REGION Network 144: Change the VG2 voltage in local
   RUNG wire#powerrail
      Contact( "STATO".controllo_setVG2 )
      wire#w1
      { S7_Templates := "SrcType := Int" } GE_Contact(in1 := "STATO".stato_VOLTAGGIO_G2, in2 := 100)
      { S7_Templates := "SrcType := Int" } LE_Contact(in1 := "STATO".stato_VOLTAGGIO_G2, in2 := 1150)
      Move(in := "STATO_TMP".tmp_adj_VG2, out1 => "STATO".stato_VOLTAGGIO_G2)
      R_Coil( "STATO".controllo_setVG2 )
   END_RUNG
   RUNG wire#w1
      { S7_Templates := "SrcType := Int" } GT_Contact(in1 := "STATO".stato_VOLTAGGIO_G2, in2 := 1150)
      Move(in := 1150, out1 => "STATO".stato_VOLTAGGIO_G2)
      R_Coil( "STATO".controllo_setVG2 )
   END_RUNG
   RUNG wire#w1
      { S7_Templates := "SrcType := Int" } LT_Contact(in1 := "STATO".stato_VOLTAGGIO_G2, in2 := 100)
      Move(in := 100, out1 => "STATO".stato_VOLTAGGIO_G2)
      R_Coil( "STATO".controllo_setVG2 )
   END_RUNG
   // the same network as SCL:
   #_w1 := "STATO".controllo_setVG2 AND ("STATO".stato_VOLTAGGIO_G2 >= 100) AND ("STATO".stato_VOLTAGGIO_G2 <= 1150);
   IF #_w1 THEN "STATO".stato_VOLTAGGIO_G2 := "STATO_TMP".tmp_adj_VG2; END_IF;
   #_w2 := "STATO".controllo_setVG2;
   IF #_w1 THEN "STATO".controllo_setVG2 := FALSE; END_IF;
   #_w3 := #_w2 AND ("STATO".stato_VOLTAGGIO_G2 > 1150);
   IF #_w3 THEN
       "STATO".stato_VOLTAGGIO_G2 := 1150;
       "STATO".controllo_setVG2 := FALSE;
   END_IF;
   #_w4 := #_w2 AND ("STATO".stato_VOLTAGGIO_G2 < 100);
   IF #_w4 THEN
       "STATO".stato_VOLTAGGIO_G2 := 100;
       "STATO".controllo_setVG2 := FALSE;
   END_IF;
END_REGION

REGION Network 145: Change the VG2 voltage in remote
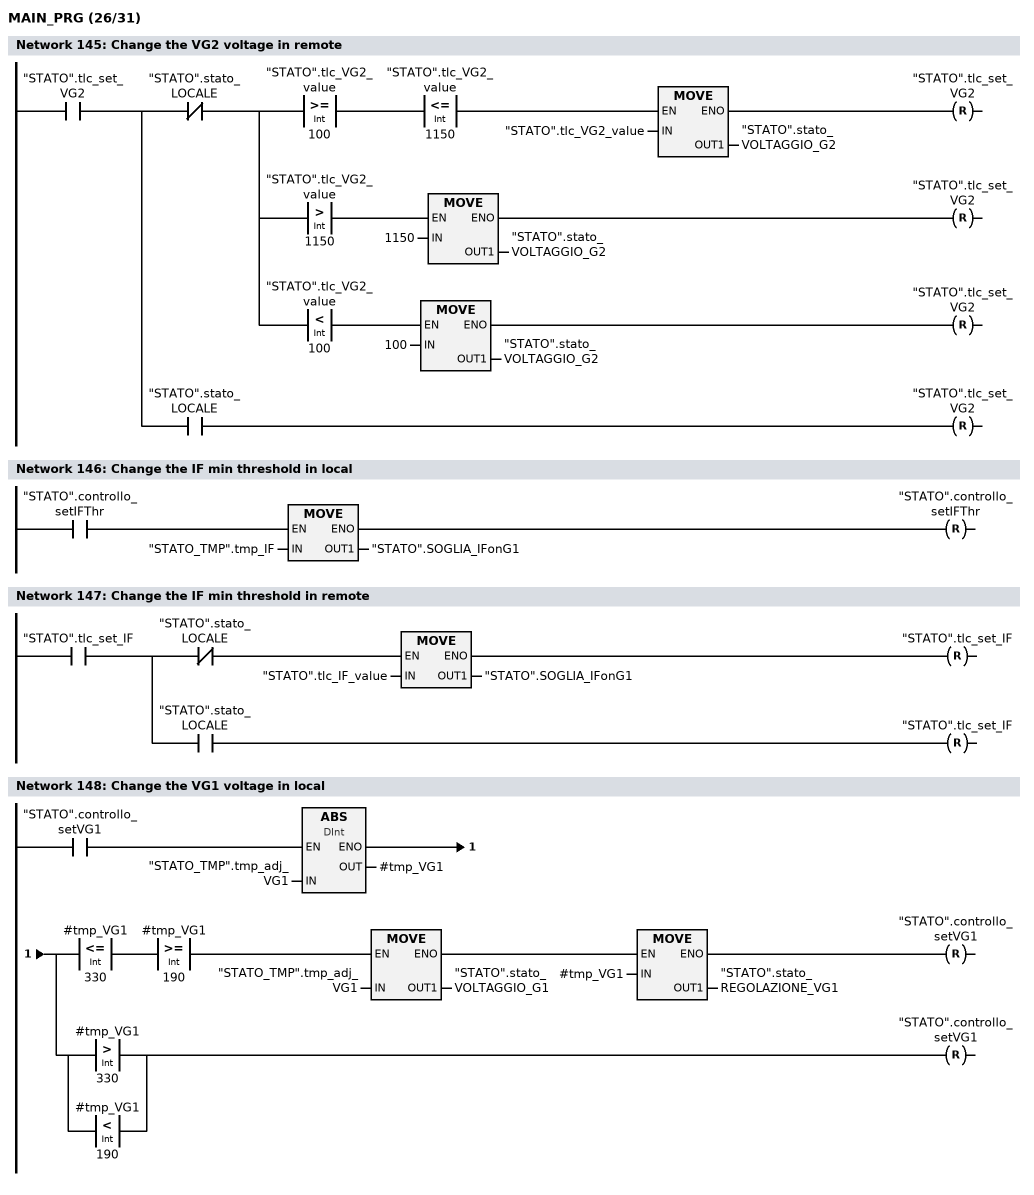
   RUNG wire#powerrail
      Contact( "STATO".tlc_set_VG2 )
      wire#w1
      I_Contact( "STATO".stato_LOCALE )
      wire#w2
      { S7_Templates := "SrcType := Int" } GE_Contact(in1 := "STATO".tlc_VG2_value, in2 := 100)
      { S7_Templates := "SrcType := Int" } LE_Contact(in1 := "STATO".tlc_VG2_value, in2 := 1150)
      Move(in := "STATO".tlc_VG2_value, out1 => "STATO".stato_VOLTAGGIO_G2)
      R_Coil( "STATO".tlc_set_VG2 )
   END_RUNG
   RUNG wire#w2
      { S7_Templates := "SrcType := Int" } GT_Contact(in1 := "STATO".tlc_VG2_value, in2 := 1150)
      Move(in := 1150, out1 => "STATO".stato_VOLTAGGIO_G2)
      R_Coil( "STATO".tlc_set_VG2 )
   END_RUNG
   RUNG wire#w2
      { S7_Templates := "SrcType := Int" } LT_Contact(in1 := "STATO".tlc_VG2_value, in2 := 100)
      Move(in := 100, out1 => "STATO".stato_VOLTAGGIO_G2)
      R_Coil( "STATO".tlc_set_VG2 )
   END_RUNG
   RUNG wire#w1
      Contact( "STATO".stato_LOCALE )
      R_Coil( "STATO".tlc_set_VG2 )
   END_RUNG
   // the same network as SCL:
   #_w1 := "STATO".tlc_set_VG2 AND NOT "STATO".stato_LOCALE;
   IF #_w1 AND ("STATO".tlc_VG2_value >= 100) AND ("STATO".tlc_VG2_value <= 1150) THEN
       "STATO".stato_VOLTAGGIO_G2 := "STATO".tlc_VG2_value;
   END_IF;
   #_w2 := "STATO".tlc_set_VG2;
   IF #_w1 AND ("STATO".tlc_VG2_value >= 100) AND ("STATO".tlc_VG2_value <= 1150) THEN
       "STATO".tlc_set_VG2 := FALSE;
   END_IF;
   IF #_w1 AND ("STATO".tlc_VG2_value > 1150) THEN
       "STATO".stato_VOLTAGGIO_G2 := 1150;
       "STATO".tlc_set_VG2 := FALSE;
   END_IF;
   IF #_w1 AND ("STATO".tlc_VG2_value < 100) THEN
       "STATO".stato_VOLTAGGIO_G2 := 100;
       "STATO".tlc_set_VG2 := FALSE;
   END_IF;
   IF #_w2 AND "STATO".stato_LOCALE THEN "STATO".tlc_set_VG2 := FALSE; END_IF;
END_REGION

REGION Network 146: Change the IF min threshold in local
   RUNG wire#powerrail
      Contact( "STATO".controllo_setIFThr )
      Move(in := "STATO_TMP".tmp_IF, out1 => "STATO".SOGLIA_IFonG1)
      R_Coil( "STATO".controllo_setIFThr )
   END_RUNG
   // the same network as SCL:
   IF "STATO".controllo_setIFThr THEN
       "STATO".SOGLIA_IFonG1 := "STATO_TMP".tmp_IF;
       "STATO".controllo_setIFThr := FALSE;
   END_IF;
END_REGION

REGION Network 147: Change the IF min threshold in remote
   RUNG wire#powerrail
      Contact( "STATO".tlc_set_IF )
      wire#w1
      I_Contact( "STATO".stato_LOCALE )
      Move(in := "STATO".tlc_IF_value, out1 => "STATO".SOGLIA_IFonG1)
      R_Coil( "STATO".tlc_set_IF )
   END_RUNG
   RUNG wire#w1
      Contact( "STATO".stato_LOCALE )
      R_Coil( "STATO".tlc_set_IF )
   END_RUNG
   // the same network as SCL:
   IF "STATO".tlc_set_IF AND NOT "STATO".stato_LOCALE THEN
       "STATO".SOGLIA_IFonG1 := "STATO".tlc_IF_value;
   END_IF;
   #_w1 := "STATO".tlc_set_IF;
   IF "STATO".tlc_set_IF AND NOT "STATO".stato_LOCALE THEN "STATO".tlc_set_IF := FALSE; END_IF;
   IF #_w1 AND "STATO".stato_LOCALE THEN "STATO".tlc_set_IF := FALSE; END_IF;
END_REGION

REGION Network 148: Change the VG1 voltage in local
   RUNG wire#powerrail
      Contact( "STATO".controllo_setVG1 )
      { S7_Templates := "SrcType := DInt" } Abs(in := "STATO_TMP".tmp_adj_VG1, out => #tmp_VG1)
      wire#w1
      { S7_Templates := "SrcType := Int" } LE_Contact(in1 := #tmp_VG1, in2 := 330)
      { S7_Templates := "SrcType := Int" } GE_Contact(in1 := #tmp_VG1, in2 := 190)
      Move(in := "STATO_TMP".tmp_adj_VG1, out1 => "STATO".stato_VOLTAGGIO_G1)
      Move(in := #tmp_VG1, out1 => "STATO".stato_REGOLAZIONE_VG1)
      R_Coil( "STATO".controllo_setVG1 )
   END_RUNG
   RUNG wire#w1
      { S7_Templates := "SrcType := Int" } GT_Contact(in1 := #tmp_VG1, in2 := 330)
      wire#w2
      R_Coil( "STATO".controllo_setVG1 )
   END_RUNG
   RUNG wire#w1
      { S7_Templates := "SrcType := Int" } LT_Contact(in1 := #tmp_VG1, in2 := 190)
   END_RUNG wire#w2
   // the same network as SCL:
   IF "STATO".controllo_setVG1 THEN #tmp_VG1 := ABS("STATO_TMP".tmp_adj_VG1); END_IF;
   IF "STATO".controllo_setVG1 AND (#tmp_VG1 <= 330) AND (#tmp_VG1 >= 190) THEN
       "STATO".stato_VOLTAGGIO_G1 := "STATO_TMP".tmp_adj_VG1;
       "STATO".stato_REGOLAZIONE_VG1 := #tmp_VG1;
   END_IF;
   #_w1 := "STATO".controllo_setVG1;
   IF "STATO".controllo_setVG1 AND (#tmp_VG1 <= 330) AND (#tmp_VG1 >= 190) THEN
       "STATO".controllo_setVG1 := FALSE;
   END_IF;
   IF #_w1 AND ((#tmp_VG1 > 330) OR (#tmp_VG1 < 190)) THEN "STATO".controllo_setVG1 := FALSE; END_IF;
END_REGION

REGION Network 149: Change the VG1 voltage in remote
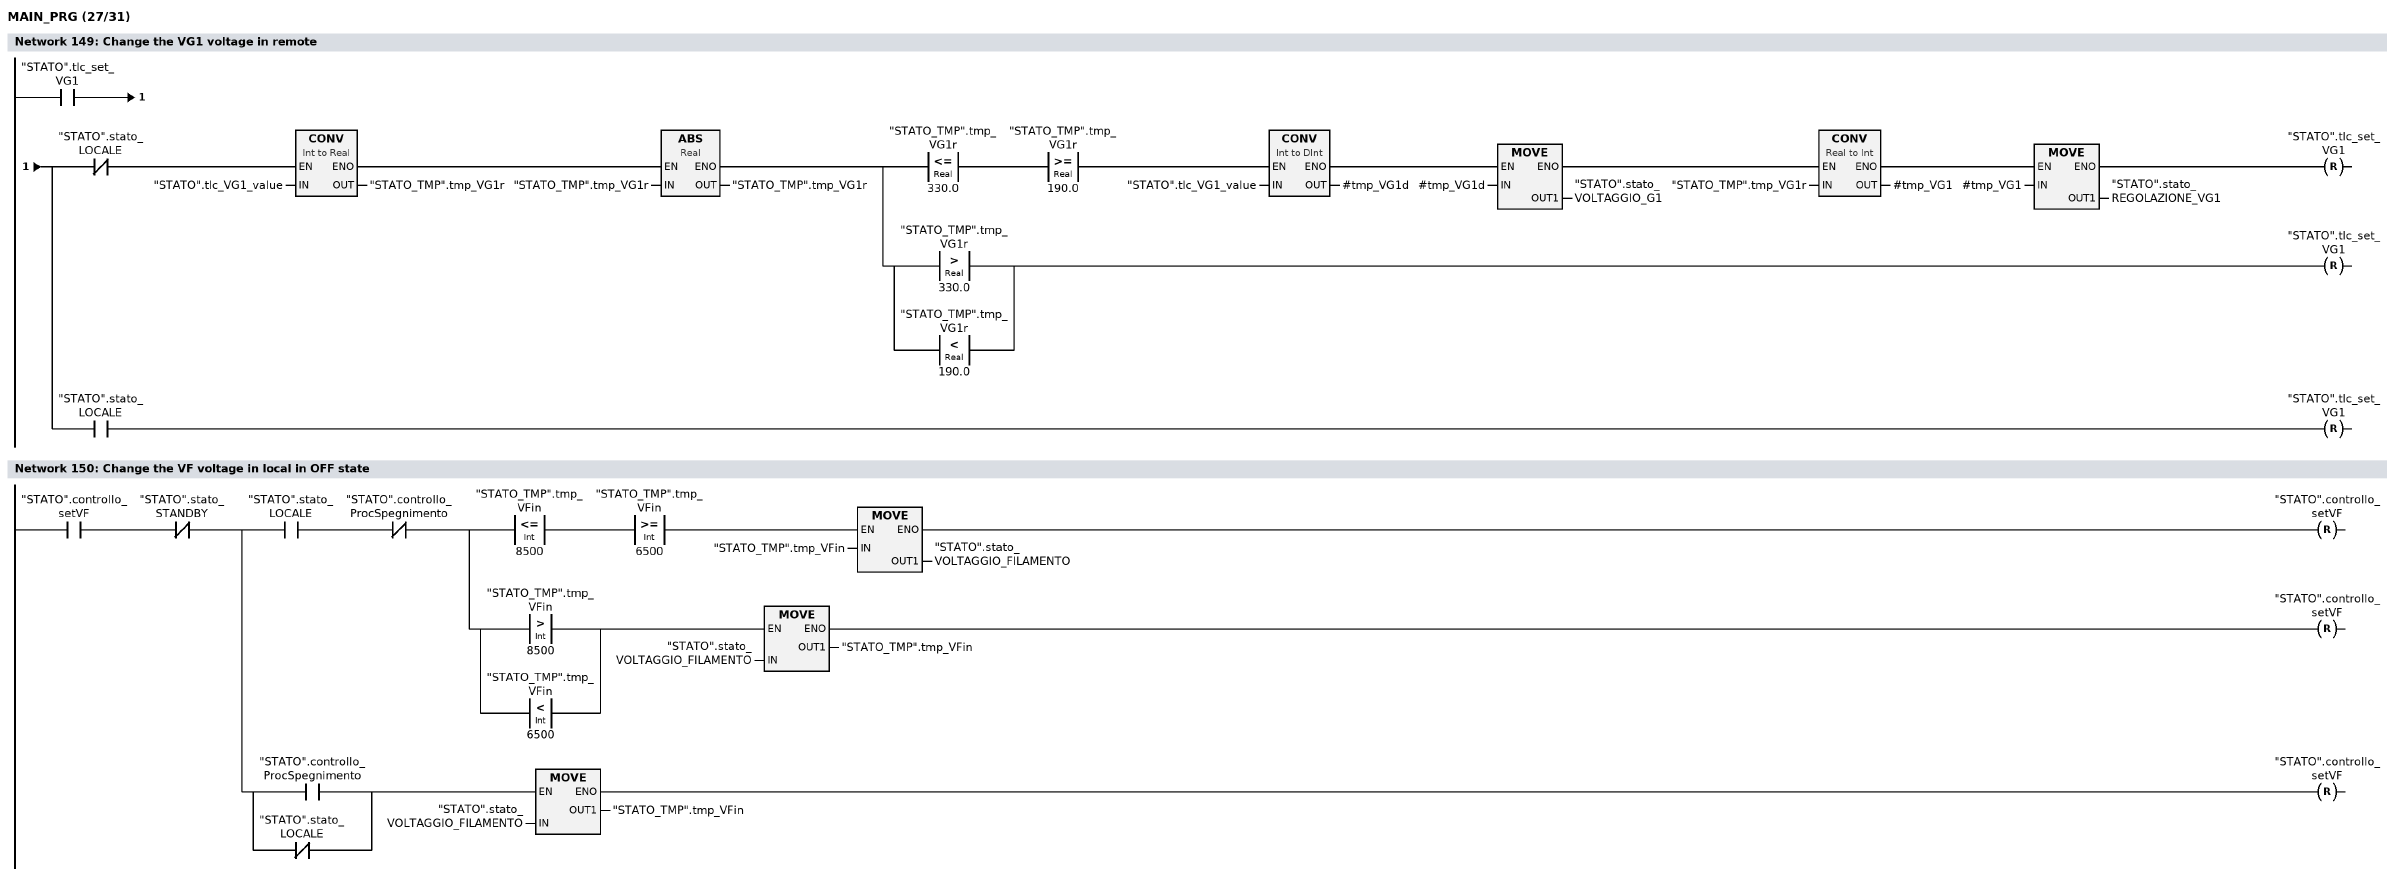
   RUNG wire#powerrail
      Contact( "STATO".tlc_set_VG1 )
      wire#w1
      I_Contact( "STATO".stato_LOCALE )
      { S7_Templates := "[SrcType := Int, DestType := Real]" } Convert(in := "STATO".tlc_VG1_value, out => "STATO_TMP".tmp_VG1r)
      { S7_Templates := "SrcType := Real" } Abs(in := "STATO_TMP".tmp_VG1r, out => "STATO_TMP".tmp_VG1r)
      wire#w2
      { S7_Templates := "SrcType := Real" } LE_Contact(in1 := "STATO_TMP".tmp_VG1r, in2 := 330.0)
      { S7_Templates := "SrcType := Real" } GE_Contact(in1 := "STATO_TMP".tmp_VG1r, in2 := 190.0)
      { S7_Templates := "[SrcType := Int, DestType := DInt]" } Convert(in := "STATO".tlc_VG1_value, out => #tmp_VG1d)
      Move(in := #tmp_VG1d, out1 => "STATO".stato_VOLTAGGIO_G1)
      { S7_Templates := "[SrcType := Real, DestType := Int]" } Convert(in := "STATO_TMP".tmp_VG1r, out => #tmp_VG1)
      Move(in := #tmp_VG1, out1 => "STATO".stato_REGOLAZIONE_VG1)
      R_Coil( "STATO".tlc_set_VG1 )
   END_RUNG
   RUNG wire#w2
      { S7_Templates := "SrcType := Real" } GT_Contact(in1 := "STATO_TMP".tmp_VG1r, in2 := 330.0)
      wire#w3
      R_Coil( "STATO".tlc_set_VG1 )
   END_RUNG
   RUNG wire#w2
      { S7_Templates := "SrcType := Real" } LT_Contact(in1 := "STATO_TMP".tmp_VG1r, in2 := 190.0)
   END_RUNG wire#w3
   RUNG wire#w1
      Contact( "STATO".stato_LOCALE )
      R_Coil( "STATO".tlc_set_VG1 )
   END_RUNG
   // the same network as SCL:
   #_w1 := "STATO".tlc_set_VG1 AND NOT "STATO".stato_LOCALE;
   IF #_w1 THEN
       "STATO_TMP".tmp_VG1r := INT_TO_REAL("STATO".tlc_VG1_value);
       "STATO_TMP".tmp_VG1r := ABS("STATO_TMP".tmp_VG1r);
   END_IF;
   IF #_w1 AND ("STATO_TMP".tmp_VG1r <= 330.0) AND ("STATO_TMP".tmp_VG1r >= 190.0) THEN
       #tmp_VG1d := INT_TO_DINT("STATO".tlc_VG1_value);
       "STATO".stato_VOLTAGGIO_G1 := #tmp_VG1d;
       #tmp_VG1 := REAL_TO_INT("STATO_TMP".tmp_VG1r);
       "STATO".stato_REGOLAZIONE_VG1 := #tmp_VG1;
   END_IF;
   #_w2 := "STATO".tlc_set_VG1;
   IF #_w1 AND ("STATO_TMP".tmp_VG1r <= 330.0) AND ("STATO_TMP".tmp_VG1r >= 190.0) THEN
       "STATO".tlc_set_VG1 := FALSE;
   END_IF;
   IF #_w1 AND (("STATO_TMP".tmp_VG1r > 330.0) OR ("STATO_TMP".tmp_VG1r < 190.0)) THEN
       "STATO".tlc_set_VG1 := FALSE;
   END_IF;
   IF #_w2 AND "STATO".stato_LOCALE THEN "STATO".tlc_set_VG1 := FALSE; END_IF;
END_REGION

REGION Network 150: Change the VF voltage in local in OFF state
   RUNG wire#powerrail
      Contact( "STATO".controllo_setVF )
      I_Contact( "STATO".stato_STANDBY )
      wire#w1
      Contact( "STATO".stato_LOCALE )
      I_Contact( "STATO".controllo_ProcSpegnimento )
      wire#w2
      { S7_Templates := "SrcType := Int" } LE_Contact(in1 := "STATO_TMP".tmp_VFin, in2 := 8500)
      { S7_Templates := "SrcType := Int" } GE_Contact(in1 := "STATO_TMP".tmp_VFin, in2 := 6500)
      Move(in := "STATO_TMP".tmp_VFin, out1 => "STATO".stato_VOLTAGGIO_FILAMENTO)
      R_Coil( "STATO".controllo_setVF )
   END_RUNG
   RUNG wire#w2
      { S7_Templates := "SrcType := Int" } GT_Contact(in1 := "STATO_TMP".tmp_VFin, in2 := 8500)
      wire#w3
      Move(in := "STATO".stato_VOLTAGGIO_FILAMENTO, out1 => "STATO_TMP".tmp_VFin)
      R_Coil( "STATO".controllo_setVF )
   END_RUNG
   RUNG wire#w2
      { S7_Templates := "SrcType := Int" } LT_Contact(in1 := "STATO_TMP".tmp_VFin, in2 := 6500)
   END_RUNG wire#w3
   RUNG wire#w1
      Contact( "STATO".controllo_ProcSpegnimento )
      wire#w4
      Move(in := "STATO".stato_VOLTAGGIO_FILAMENTO, out1 => "STATO_TMP".tmp_VFin)
      R_Coil( "STATO".controllo_setVF )
   END_RUNG
   RUNG wire#w1
      I_Contact( "STATO".stato_LOCALE )
   END_RUNG wire#w4
   // the same network as SCL:
   #_w1 := "STATO".controllo_setVF AND NOT "STATO".stato_STANDBY;
   #_w2 := #_w1 AND "STATO".stato_LOCALE AND NOT "STATO".controllo_ProcSpegnimento;
   IF #_w2 AND ("STATO_TMP".tmp_VFin <= 8500) AND ("STATO_TMP".tmp_VFin >= 6500) THEN
       "STATO".stato_VOLTAGGIO_FILAMENTO := "STATO_TMP".tmp_VFin;
       "STATO".controllo_setVF := FALSE;
   END_IF;
   #_w3 := #_w2 AND (("STATO_TMP".tmp_VFin > 8500) OR ("STATO_TMP".tmp_VFin < 6500));
   IF #_w3 THEN
       "STATO_TMP".tmp_VFin := "STATO".stato_VOLTAGGIO_FILAMENTO;
       "STATO".controllo_setVF := FALSE;
   END_IF;
   IF #_w1 AND ("STATO".controllo_ProcSpegnimento OR NOT "STATO".stato_LOCALE) THEN
       "STATO_TMP".tmp_VFin := "STATO".stato_VOLTAGGIO_FILAMENTO;
       "STATO".controllo_setVF := FALSE;
   END_IF;
END_REGION

REGION Network 151: Change the VF voltage in local during operation
   // change the filament voltage in 100mV step
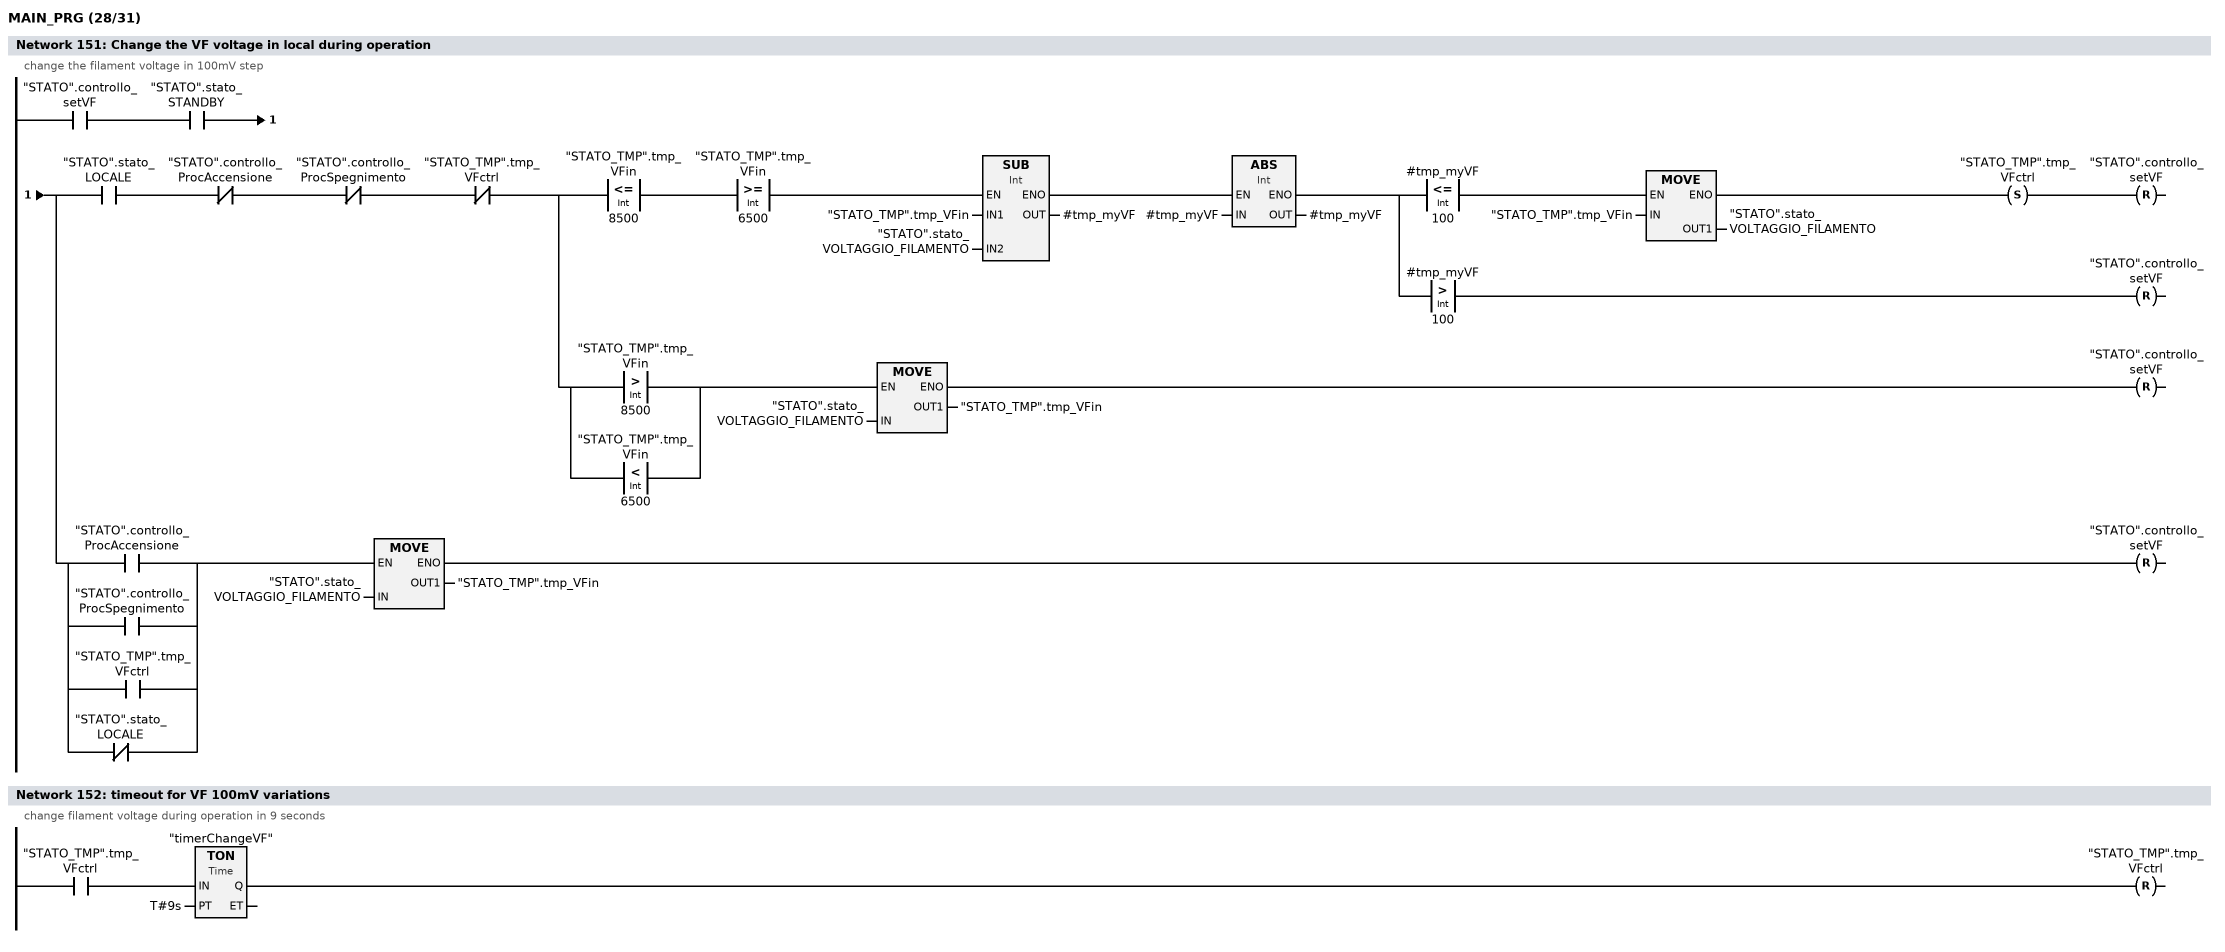
   RUNG wire#powerrail
      Contact( "STATO".controllo_setVF )
      Contact( "STATO".stato_STANDBY )
      wire#w1
      Contact( "STATO".stato_LOCALE )
      I_Contact( "STATO".controllo_ProcAccensione )
      I_Contact( "STATO".controllo_ProcSpegnimento )
      I_Contact( "STATO_TMP".tmp_VFctrl )
      wire#w2
      { S7_Templates := "SrcType := Int" } LE_Contact(in1 := "STATO_TMP".tmp_VFin, in2 := 8500)
      { S7_Templates := "SrcType := Int" } GE_Contact(in1 := "STATO_TMP".tmp_VFin, in2 := 6500)
      { S7_Templates := "SrcType := Int" } Sub(in1 := "STATO_TMP".tmp_VFin, in2 := "STATO".stato_VOLTAGGIO_FILAMENTO, out => #tmp_myVF)
      { S7_Templates := "SrcType := Int" } Abs(in := #tmp_myVF, out => #tmp_myVF)
      wire#w3
      { S7_Templates := "SrcType := Int" } LE_Contact(in1 := #tmp_myVF, in2 := 100)
      Move(in := "STATO_TMP".tmp_VFin, out1 => "STATO".stato_VOLTAGGIO_FILAMENTO)
      S_Coil( "STATO_TMP".tmp_VFctrl )
      R_Coil( "STATO".controllo_setVF )
   END_RUNG
   RUNG wire#w3
      { S7_Templates := "SrcType := Int" } GT_Contact(in1 := #tmp_myVF, in2 := 100)
      R_Coil( "STATO".controllo_setVF )
   END_RUNG
   RUNG wire#w2
      { S7_Templates := "SrcType := Int" } GT_Contact(in1 := "STATO_TMP".tmp_VFin, in2 := 8500)
      wire#w4
      Move(in := "STATO".stato_VOLTAGGIO_FILAMENTO, out1 => "STATO_TMP".tmp_VFin)
      R_Coil( "STATO".controllo_setVF )
   END_RUNG
   RUNG wire#w2
      { S7_Templates := "SrcType := Int" } LT_Contact(in1 := "STATO_TMP".tmp_VFin, in2 := 6500)
   END_RUNG wire#w4
   RUNG wire#w1
      Contact( "STATO".controllo_ProcAccensione )
      wire#w5
      Move(in := "STATO".stato_VOLTAGGIO_FILAMENTO, out1 => "STATO_TMP".tmp_VFin)
      R_Coil( "STATO".controllo_setVF )
   END_RUNG
   RUNG wire#w1
      Contact( "STATO".controllo_ProcSpegnimento )
   END_RUNG wire#w5
   RUNG wire#w1
      Contact( "STATO_TMP".tmp_VFctrl )
   END_RUNG wire#w5
   RUNG wire#w1
      I_Contact( "STATO".stato_LOCALE )
   END_RUNG wire#w5
   // the same network as SCL:
   #_w1 := "STATO".controllo_setVF AND "STATO".stato_STANDBY;
   #_w2 := #_w1 AND "STATO".stato_LOCALE AND NOT "STATO".controllo_ProcAccensione AND NOT "STATO".controllo_ProcSpegnimento AND NOT "STATO_TMP".tmp_VFctrl;
   #_w3 := #_w2 AND ("STATO_TMP".tmp_VFin <= 8500) AND ("STATO_TMP".tmp_VFin >= 6500);
   IF #_w3 THEN
       #tmp_myVF := "STATO_TMP".tmp_VFin - "STATO".stato_VOLTAGGIO_FILAMENTO;
       #tmp_myVF := ABS(#tmp_myVF);
   END_IF;
   IF #_w3 AND (#tmp_myVF <= 100) THEN
       "STATO".stato_VOLTAGGIO_FILAMENTO := "STATO_TMP".tmp_VFin;
       "STATO_TMP".tmp_VFctrl := TRUE;
       "STATO".controllo_setVF := FALSE;
   END_IF;
   IF #_w3 AND (#tmp_myVF > 100) THEN "STATO".controllo_setVF := FALSE; END_IF;
   #_w4 := #_w2 AND (("STATO_TMP".tmp_VFin > 8500) OR ("STATO_TMP".tmp_VFin < 6500));
   IF #_w4 THEN
       "STATO_TMP".tmp_VFin := "STATO".stato_VOLTAGGIO_FILAMENTO;
       "STATO".controllo_setVF := FALSE;
   END_IF;
   IF #_w1 AND ("STATO".controllo_ProcAccensione OR "STATO".controllo_ProcSpegnimento OR "STATO_TMP".tmp_VFctrl OR NOT "STATO".stato_LOCALE) THEN
       "STATO_TMP".tmp_VFin := "STATO".stato_VOLTAGGIO_FILAMENTO;
       "STATO".controllo_setVF := FALSE;
   END_IF;
END_REGION

REGION Network 152: timeout for VF 100mV variations
   // change filament voltage during operation in 9 seconds
   "timerChangeVF".TON(IN := "STATO_TMP".tmp_VFctrl, PT := T#9s);
   IF "timerChangeVF".Q THEN "STATO_TMP".tmp_VFctrl := FALSE; END_IF;
END_REGION

REGION Network 153: Change the VF voltage in remote
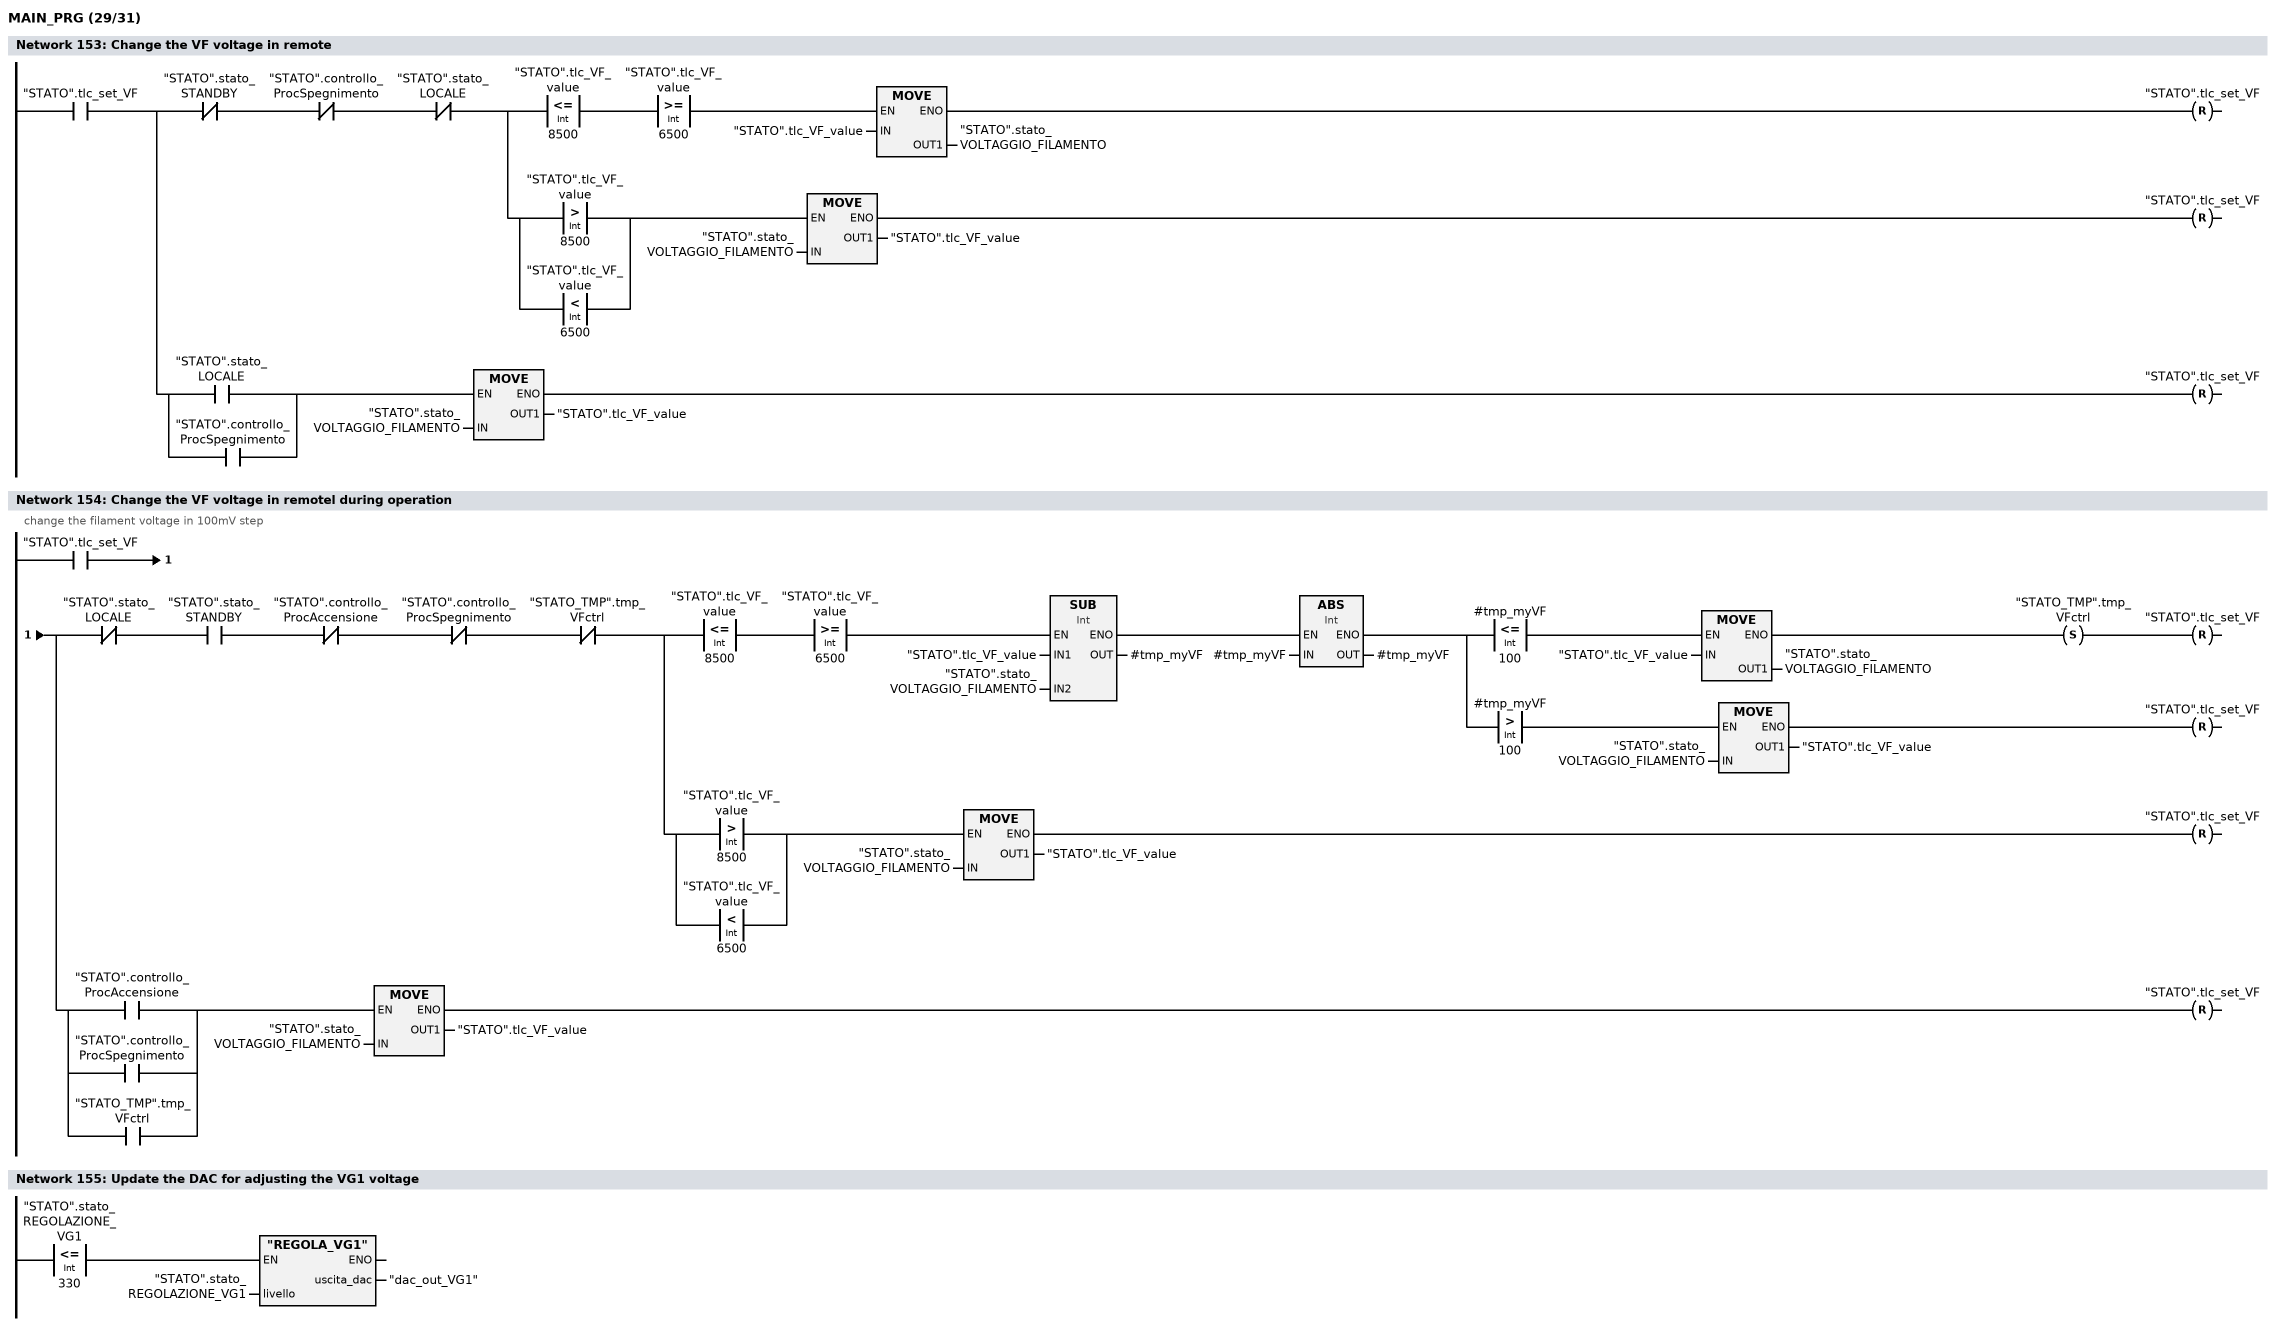
   RUNG wire#powerrail
      Contact( "STATO".tlc_set_VF )
      wire#w1
      I_Contact( "STATO".stato_STANDBY )
      I_Contact( "STATO".controllo_ProcSpegnimento )
      I_Contact( "STATO".stato_LOCALE )
      wire#w2
      { S7_Templates := "SrcType := Int" } LE_Contact(in1 := "STATO".tlc_VF_value, in2 := 8500)
      { S7_Templates := "SrcType := Int" } GE_Contact(in1 := "STATO".tlc_VF_value, in2 := 6500)
      Move(in := "STATO".tlc_VF_value, out1 => "STATO".stato_VOLTAGGIO_FILAMENTO)
      R_Coil( "STATO".tlc_set_VF )
   END_RUNG
   RUNG wire#w2
      { S7_Templates := "SrcType := Int" } GT_Contact(in1 := "STATO".tlc_VF_value, in2 := 8500)
      wire#w3
      Move(in := "STATO".stato_VOLTAGGIO_FILAMENTO, out1 => "STATO".tlc_VF_value)
      R_Coil( "STATO".tlc_set_VF )
   END_RUNG
   RUNG wire#w2
      { S7_Templates := "SrcType := Int" } LT_Contact(in1 := "STATO".tlc_VF_value, in2 := 6500)
   END_RUNG wire#w3
   RUNG wire#w1
      Contact( "STATO".stato_LOCALE )
      wire#w4
      Move(in := "STATO".stato_VOLTAGGIO_FILAMENTO, out1 => "STATO".tlc_VF_value)
      R_Coil( "STATO".tlc_set_VF )
   END_RUNG
   RUNG wire#w1
      Contact( "STATO".controllo_ProcSpegnimento )
   END_RUNG wire#w4
   // the same network as SCL:
   #_w1 := "STATO".tlc_set_VF AND NOT "STATO".stato_STANDBY AND NOT "STATO".controllo_ProcSpegnimento AND NOT "STATO".stato_LOCALE;
   IF #_w1 AND ("STATO".tlc_VF_value <= 8500) AND ("STATO".tlc_VF_value >= 6500) THEN
       "STATO".stato_VOLTAGGIO_FILAMENTO := "STATO".tlc_VF_value;
   END_IF;
   #_w2 := "STATO".tlc_set_VF;
   IF #_w1 AND ("STATO".tlc_VF_value <= 8500) AND ("STATO".tlc_VF_value >= 6500) THEN
       "STATO".tlc_set_VF := FALSE;
   END_IF;
   #_w3 := #_w1 AND (("STATO".tlc_VF_value > 8500) OR ("STATO".tlc_VF_value < 6500));
   IF #_w3 THEN
       "STATO".tlc_VF_value := "STATO".stato_VOLTAGGIO_FILAMENTO;
       "STATO".tlc_set_VF := FALSE;
   END_IF;
   IF #_w2 AND ("STATO".stato_LOCALE OR "STATO".controllo_ProcSpegnimento) THEN
       "STATO".tlc_VF_value := "STATO".stato_VOLTAGGIO_FILAMENTO;
       "STATO".tlc_set_VF := FALSE;
   END_IF;
END_REGION

REGION Network 154: Change the VF voltage in remotel during operation
   // change the filament voltage in 100mV step
   RUNG wire#powerrail
      Contact( "STATO".tlc_set_VF )
      wire#w1
      I_Contact( "STATO".stato_LOCALE )
      Contact( "STATO".stato_STANDBY )
      I_Contact( "STATO".controllo_ProcAccensione )
      I_Contact( "STATO".controllo_ProcSpegnimento )
      I_Contact( "STATO_TMP".tmp_VFctrl )
      wire#w2
      { S7_Templates := "SrcType := Int" } LE_Contact(in1 := "STATO".tlc_VF_value, in2 := 8500)
      { S7_Templates := "SrcType := Int" } GE_Contact(in1 := "STATO".tlc_VF_value, in2 := 6500)
      { S7_Templates := "SrcType := Int" } Sub(in1 := "STATO".tlc_VF_value, in2 := "STATO".stato_VOLTAGGIO_FILAMENTO, out => #tmp_myVF)
      { S7_Templates := "SrcType := Int" } Abs(in := #tmp_myVF, out => #tmp_myVF)
      wire#w3
      { S7_Templates := "SrcType := Int" } LE_Contact(in1 := #tmp_myVF, in2 := 100)
      Move(in := "STATO".tlc_VF_value, out1 => "STATO".stato_VOLTAGGIO_FILAMENTO)
      S_Coil( "STATO_TMP".tmp_VFctrl )
      R_Coil( "STATO".tlc_set_VF )
   END_RUNG
   RUNG wire#w3
      { S7_Templates := "SrcType := Int" } GT_Contact(in1 := #tmp_myVF, in2 := 100)
      Move(in := "STATO".stato_VOLTAGGIO_FILAMENTO, out1 => "STATO".tlc_VF_value)
      R_Coil( "STATO".tlc_set_VF )
   END_RUNG
   RUNG wire#w2
      { S7_Templates := "SrcType := Int" } GT_Contact(in1 := "STATO".tlc_VF_value, in2 := 8500)
      wire#w4
      Move(in := "STATO".stato_VOLTAGGIO_FILAMENTO, out1 => "STATO".tlc_VF_value)
      R_Coil( "STATO".tlc_set_VF )
   END_RUNG
   RUNG wire#w2
      { S7_Templates := "SrcType := Int" } LT_Contact(in1 := "STATO".tlc_VF_value, in2 := 6500)
   END_RUNG wire#w4
   RUNG wire#w1
      Contact( "STATO".controllo_ProcAccensione )
      wire#w5
      Move(in := "STATO".stato_VOLTAGGIO_FILAMENTO, out1 => "STATO".tlc_VF_value)
      R_Coil( "STATO".tlc_set_VF )
   END_RUNG
   RUNG wire#w1
      Contact( "STATO".controllo_ProcSpegnimento )
   END_RUNG wire#w5
   RUNG wire#w1
      Contact( "STATO_TMP".tmp_VFctrl )
   END_RUNG wire#w5
   // the same network as SCL:
   #_w1 := "STATO".tlc_set_VF AND NOT "STATO".stato_LOCALE AND "STATO".stato_STANDBY AND NOT "STATO".controllo_ProcAccensione AND NOT "STATO".controllo_ProcSpegnimento AND NOT "STATO_TMP".tmp_VFctrl;
   #_w2 := #_w1 AND ("STATO".tlc_VF_value <= 8500) AND ("STATO".tlc_VF_value >= 6500);
   IF #_w2 THEN
       #tmp_myVF := "STATO".tlc_VF_value - "STATO".stato_VOLTAGGIO_FILAMENTO;
       #tmp_myVF := ABS(#tmp_myVF);
   END_IF;
   IF #_w2 AND (#tmp_myVF <= 100) THEN
       "STATO".stato_VOLTAGGIO_FILAMENTO := "STATO".tlc_VF_value;
       "STATO_TMP".tmp_VFctrl := TRUE;
   END_IF;
   #_w3 := "STATO".tlc_set_VF;
   IF #_w2 AND (#tmp_myVF <= 100) THEN "STATO".tlc_set_VF := FALSE; END_IF;
   IF #_w2 AND (#tmp_myVF > 100) THEN
       "STATO".tlc_VF_value := "STATO".stato_VOLTAGGIO_FILAMENTO;
       "STATO".tlc_set_VF := FALSE;
   END_IF;
   #_w4 := #_w1 AND (("STATO".tlc_VF_value > 8500) OR ("STATO".tlc_VF_value < 6500));
   IF #_w4 THEN
       "STATO".tlc_VF_value := "STATO".stato_VOLTAGGIO_FILAMENTO;
       "STATO".tlc_set_VF := FALSE;
   END_IF;
   IF #_w3 AND ("STATO".controllo_ProcAccensione OR "STATO".controllo_ProcSpegnimento OR "STATO_TMP".tmp_VFctrl) THEN
       "STATO".tlc_VF_value := "STATO".stato_VOLTAGGIO_FILAMENTO;
       "STATO".tlc_set_VF := FALSE;
   END_IF;
END_REGION

REGION Network 155: Update the DAC for adjusting the VG1 voltage
   RUNG wire#powerrail
      { S7_Templates := "SrcType := Int" } LE_Contact(in1 := "STATO".stato_REGOLAZIONE_VG1, in2 := 330)
      "REGOLA_VG1"(livello := "STATO".stato_REGOLAZIONE_VG1, uscita_dac => "dac_out_VG1")
   END_RUNG
   // the same network as SCL:
   IF "STATO".stato_REGOLAZIONE_VG1 <= 330 THEN
       "REGOLA_VG1"(livello := "STATO".stato_REGOLAZIONE_VG1, uscita_dac => "dac_out_VG1");
   END_IF;
END_REGION

REGION Network 156: Update the DAC for adjusting the VG1 voltage
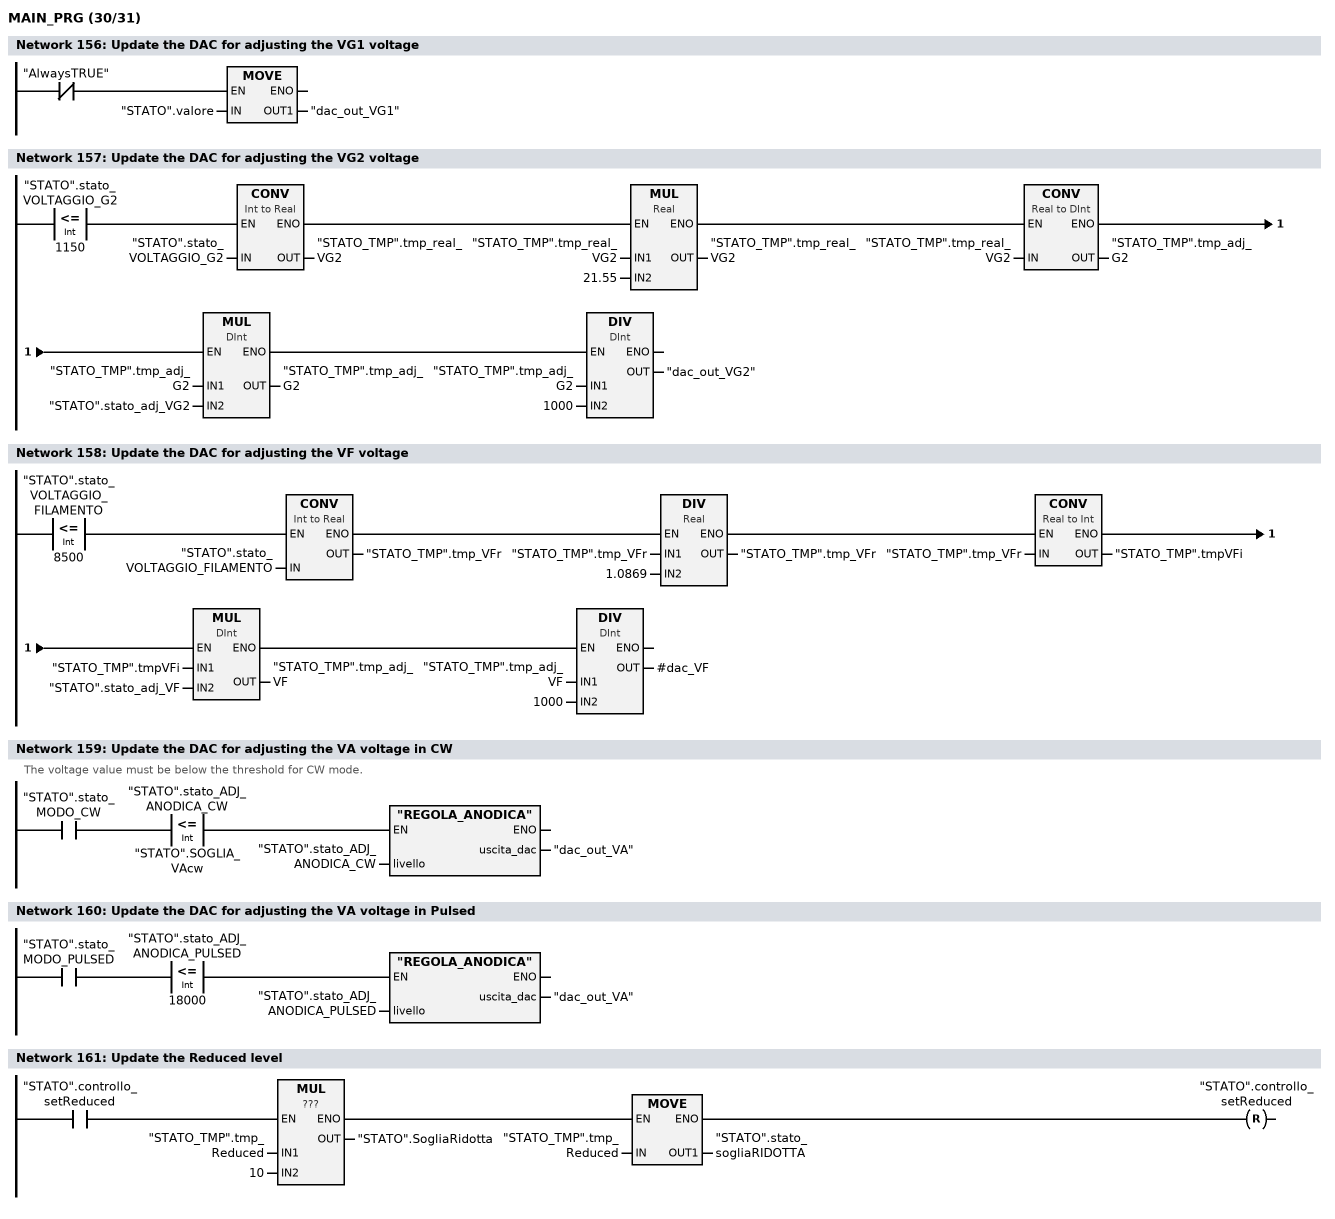
   RUNG wire#powerrail
      I_Contact( "AlwaysTRUE" )
      Move(in := "STATO".valore, out1 => "dac_out_VG1")
   END_RUNG
   // the same network as SCL:
   IF NOT "AlwaysTRUE" THEN "dac_out_VG1" := "STATO".valore; END_IF;
END_REGION
